   2804: 'Spare_Fault_2804', class No Acknowledgement, trigger "DB302_HMI_Faults_Carrier43_Faults_3" bit 3
   2805: 'Spare_Fault_2805', class No Acknowledgement, trigger "DB302_HMI_Faults_Carrier43_Faults_3" bit 4
   2806: 'Spare_Fault_2806', class No Acknowledgement, trigger "DB302_HMI_Faults_Carrier43_Faults_3" bit 5
   2807: 'Spare_Fault_2807', class No Acknowledgement, trigger "DB302_HMI_Faults_Carrier43_Faults_3" bit 6
   2808: 'Spare_Fault_2808', class No Acknowledgement, trigger "DB302_HMI_Faults_Carrier43_Faults_3" bit 7
   2809: 'Spare_Fault_2809', class No Acknowledgement, trigger "DB302_HMI_Faults_Carrier43_Faults_3" bit 8
   2810: 'Spare_Fault_2810', class No Acknowledgement, trigger "DB302_HMI_Faults_Carrier43_Faults_3" bit 9
   2811: 'Spare_Fault_2811', class No Acknowledgement, trigger "DB302_HMI_Faults_Carrier43_Faults_3" bit 10
   2812: 'Spare_Fault_2812', class No Acknowledgement, trigger "DB302_HMI_Faults_Carrier43_Faults_3" bit 11
   2813: 'Spare_Fault_2813', class No Acknowledgement, trigger "DB302_HMI_Faults_Carrier43_Faults_3" bit 12
   2814: 'Spare_Fault_2814', class No Acknowledgement, trigger "DB302_HMI_Faults_Carrier43_Faults_3" bit 13
   2815: 'Spare_Fault_2815', class No Acknowledgement, trigger "DB302_HMI_Faults_Carrier43_Faults_3" bit 14
   2816: 'Spare_Fault_2816', class No Acknowledgement, trigger "DB302_HMI_Faults_Carrier43_Faults_3" bit 15
   2817: 'Carrier 44 Disconnect Open Power Fault DI11.0', class No Acknowledgement, trigger "DB302_HMI_Faults_Carrier44_Faults_0" bit 0
   2818: 'Carrier 44 Drive Profinet Comm Fault', class No Acknowledgement, trigger "DB302_HMI_Faults_Carrier44_Faults_0" bit 1
   2819: 'Carrier 44 Production Stop Not Reset', class No Acknowledgement, trigger "DB302_HMI_Faults_Carrier44_Faults_0" bit 2
   2820: 'Carrier 44 CB02122 Tripped', class No Acknowledgement, trigger "DB302_HMI_Faults_Carrier44_Faults_0" bit 3
   2821: 'Carrier 44 CB02123 Tripped', class No Acknowledgement, trigger "DB302_HMI_Faults_Carrier44_Faults_0" bit 4
   2822: 'Carrier 44 AUX1 CB Tripped', class No Acknowledgement, trigger "DB302_HMI_Faults_Carrier44_Faults_0" bit 5
   2823: 'Carrier 44 AUX2 CB Tripped', class No Acknowledgement, trigger "DB302_HMI_Faults_Carrier44_Faults_0" bit 6
   2824: 'Carrier 44 PLC Not Communicating', class No Acknowledgement, trigger "DB302_HMI_Faults_Carrier44_Faults_0" bit 7
   2825: 'Carrier 44 Safe Input Card Fault', class No Acknowledgement, trigger "DB302_HMI_Faults_Carrier44_Faults_0" bit 8
   2826: 'Carrier 44 Safe Output Card Fault', class No Acknowledgement, trigger "DB302_HMI_Faults_Carrier44_Faults_0" bit 9
   2827: 'Carrier 44 Standard Input Card Fault', class No Acknowledgement, trigger "DB302_HMI_Faults_Carrier44_Faults_0" bit 10
   2828: 'Carrier 44 Standard Output Card Fault', class No Acknowledgement, trigger "DB302_HMI_Faults_Carrier44_Faults_0" bit 11
   2829: 'Carrier 44 Encoder Position Fault', class No Acknowledgement, trigger "DB302_HMI_Faults_Carrier44_Faults_0" bit 12
   2830: 'Carrier 44 Encoder Internal Error', class No Acknowledgement, trigger "DB302_HMI_Faults_Carrier44_Faults_0" bit 13
   2831: 'Carrier 44 Encoder Comm Fault', class No Acknowledgement, trigger "DB302_HMI_Faults_Carrier44_Faults_0" bit 14
   2832: 'Carrier 44 HMI Comm Fault', class No Acknowledgement, trigger "DB302_HMI_Faults_Carrier44_Faults_0" bit 15
   2833: 'Carrier 44 Crash Detection Fault', class No Acknowledgement, trigger "DB302_HMI_Faults_Carrier44_Faults_1" bit 0
   2834: 'Carrier 44 Carrier Number Invalid', class No Acknowledgement, trigger "DB302_HMI_Faults_Carrier44_Faults_1" bit 1
   2835: 'Carrier 44 Drive: PROFINET configuration error', class No Acknowledgement, trigger "DB302_HMI_Faults_Carrier44_Faults_1" bit 2
   2836: 'Carrier 44 Drive: Error internal communications', class No Acknowledgement, trigger "DB302_HMI_Faults_Carrier44_Faults_1" bit 3
   2837: 'Carrier 44 Drive: Motor overtemperature', class No Acknowledgement, trigger "DB302_HMI_Faults_Carrier44_Faults_1" bit 4
   2838: 'Carrier 44 Drive: Motor overcurrent', class No Acknowledgement, trigger "DB302_HMI_Faults_Carrier44_Faults_1" bit 5
   2839: 'Carrier 44 Drive: Infeed or power unit not ready', class No Acknowledgement, trigger "DB302_HMI_Faults_Carrier44_Faults_1" bit 6
   2840: 'Carrier 44 Drive: Short-circuit/ground fault detected', class No Acknowledgement, trigger "DB302_HMI_Faults_Carrier44_Faults_1" bit 7
   2841: 'Carrier 44 Drive: PROFINET Setpoint timeout', class No Acknowledgement, trigger "DB302_HMI_Faults_Carrier44_Faults_1" bit 8
   2842: 'Carrier 44 Power unit: Overcurrent', class No Acknowledgement, trigger "DB302_HMI_Faults_Carrier44_Faults_1" bit 9
   2843: 'Carrier 44 Power unit: DC link voltage overvoltage', class No Acknowledgement, trigger "DB302_HMI_Faults_Carrier44_Faults_1" bit 10
   2844: 'Carrier 44 Power unit: DC link voltage undervoltage', class No Acknowledgement, trigger "DB302_HMI_Faults_Carrier44_Faults_1" bit 11
   2845: 'Carrier 44 Power unit: Line phase failure in main circuit', class No Acknowledgement, trigger "DB302_HMI_Faults_Carrier44_Faults_1" bit 12
   2846: 'Carrier 44 Power unit: Phase failure motor cable', class No Acknowledgement, trigger "DB302_HMI_Faults_Carrier44_Faults_1" bit 13
   2847: 'Carrier 44 Power unit: Ground fault', class No Acknowledgement, trigger "DB302_HMI_Faults_Carrier44_Faults_1" bit 14
   2848: 'Spare_Fault_2848', class No Acknowledgement, trigger "DB302_HMI_Faults_Carrier44_Faults_1" bit 15
   2849: 'Carrier 44 Motion Off Fault', class No Acknowledgement, trigger "DB302_HMI_Faults_Carrier44_Faults_2" bit 0
   2850: 'Carrier 44 Motion On Fault', class No Acknowledgement, trigger "DB302_HMI_Faults_Carrier44_Faults_2" bit 1
   2851: 'Carrier 44 Spacing Fault', class No Acknowledgement, trigger "DB302_HMI_Faults_Carrier44_Faults_2" bit 2
   2852: 'Carrier 44 Duplicate Carrier Number Fault', class No Acknowledgement, trigger "DB302_HMI_Faults_Carrier44_Faults_2" bit 3
   2853: 'Spare_Fault_2853', class No Acknowledgement, trigger "DB302_HMI_Faults_Carrier44_Faults_2" bit 4
   2854: 'Spare_Fault_2854', class No Acknowledgement, trigger "DB302_HMI_Faults_Carrier44_Faults_2" bit 5
   2855: 'Spare_Fault_2855', class No Acknowledgement, trigger "DB302_HMI_Faults_Carrier44_Faults_2" bit 6
   2856: 'Spare_Fault_2856', class No Acknowledgement, trigger "DB302_HMI_Faults_Carrier44_Faults_2" bit 7
   2857: 'Spare_Fault_2857', class No Acknowledgement, trigger "DB302_HMI_Faults_Carrier44_Faults_2" bit 8
   2858: 'Spare_Fault_2858', class No Acknowledgement, trigger "DB302_HMI_Faults_Carrier44_Faults_2" bit 9
   2859: 'Spare_Fault_2859', class No Acknowledgement, trigger "DB302_HMI_Faults_Carrier44_Faults_2" bit 10
   2860: 'Spare_Fault_2860', class No Acknowledgement, trigger "DB302_HMI_Faults_Carrier44_Faults_2" bit 11
   2861: 'Spare_Fault_2861', class No Acknowledgement, trigger "DB302_HMI_Faults_Carrier44_Faults_2" bit 12
   2862: 'Spare_Fault_2862', class No Acknowledgement, trigger "DB302_HMI_Faults_Carrier44_Faults_2" bit 13
   2863: 'Spare_Fault_2863', class No Acknowledgement, trigger "DB302_HMI_Faults_Carrier44_Faults_2" bit 14
   2864: 'Spare_Fault_2864', class No Acknowledgement, trigger "DB302_HMI_Faults_Carrier44_Faults_2" bit 15
   2865: 'Spare_Fault_2865', class No Acknowledgement, trigger "DB302_HMI_Faults_Carrier44_Faults_3" bit 0
   2866: 'Spare_Fault_2866', class No Acknowledgement, trigger "DB302_HMI_Faults_Carrier44_Faults_3" bit 1
   2867: 'Spare_Fault_2867', class No Acknowledgement, trigger "DB302_HMI_Faults_Carrier44_Faults_3" bit 2
   2868: 'Spare_Fault_2868', class No Acknowledgement, trigger "DB302_HMI_Faults_Carrier44_Faults_3" bit 3
   2869: 'Spare_Fault_2869', class No Acknowledgement, trigger "DB302_HMI_Faults_Carrier44_Faults_3" bit 4
   2870: 'Spare_Fault_2870', class No Acknowledgement, trigger "DB302_HMI_Faults_Carrier44_Faults_3" bit 5
   2871: 'Spare_Fault_2871', class No Acknowledgement, trigger "DB302_HMI_Faults_Carrier44_Faults_3" bit 6
   2872: 'Spare_Fault_2872', class No Acknowledgement, trigger "DB302_HMI_Faults_Carrier44_Faults_3" bit 7
   2873: 'Spare_Fault_2873', class No Acknowledgement, trigger "DB302_HMI_Faults_Carrier44_Faults_3" bit 8
   2874: 'Spare_Fault_2874', class No Acknowledgement, trigger "DB302_HMI_Faults_Carrier44_Faults_3" bit 9
   2875: 'Spare_Fault_2875', class No Acknowledgement, trigger "DB302_HMI_Faults_Carrier44_Faults_3" bit 10
   2876: 'Spare_Fault_2876', class No Acknowledgement, trigger "DB302_HMI_Faults_Carrier44_Faults_3" bit 11
   2877: 'Spare_Fault_2877', class No Acknowledgement, trigger "DB302_HMI_Faults_Carrier44_Faults_3" bit 12
   2878: 'Spare_Fault_2878', class No Acknowledgement, trigger "DB302_HMI_Faults_Carrier44_Faults_3" bit 13
   2879: 'Spare_Fault_2879', class No Acknowledgement, trigger "DB302_HMI_Faults_Carrier44_Faults_3" bit 14
   2880: 'Spare_Fault_2880', class No Acknowledgement, trigger "DB302_HMI_Faults_Carrier44_Faults_3" bit 15
   2881: 'Carrier 45 Disconnect Open Power Fault DI11.0', class No Acknowledgement, trigger "DB302_HMI_Faults_Carrier45_Faults_0" bit 0
   2882: 'Carrier 45 Drive Profinet Comm Fault', class No Acknowledgement, trigger "DB302_HMI_Faults_Carrier45_Faults_0" bit 1
   2883: 'Carrier 45 Production Stop Not Reset', class No Acknowledgement, trigger "DB302_HMI_Faults_Carrier45_Faults_0" bit 2
   2884: 'Carrier 45 CB02122 Tripped', class No Acknowledgement, trigger "DB302_HMI_Faults_Carrier45_Faults_0" bit 3
   2885: 'Carrier 45 CB02123 Tripped', class No Acknowledgement, trigger "DB302_HMI_Faults_Carrier45_Faults_0" bit 4
   2886: 'Carrier 45 AUX1 CB Tripped', class No Acknowledgement, trigger "DB302_HMI_Faults_Carrier45_Faults_0" bit 5
   2887: 'Carrier 45 AUX2 CB Tripped', class No Acknowledgement, trigger "DB302_HMI_Faults_Carrier45_Faults_0" bit 6
   2888: 'Carrier 45 PLC Not Communicating', class No Acknowledgement, trigger "DB302_HMI_Faults_Carrier45_Faults_0" bit 7
   2889: 'Carrier 45 Safe Input Card Fault', class No Acknowledgement, trigger "DB302_HMI_Faults_Carrier45_Faults_0" bit 8
   2890: 'Carrier 45 Safe Output Card Fault', class No Acknowledgement, trigger "DB302_HMI_Faults_Carrier45_Faults_0" bit 9
   2891: 'Carrier 45 Standard Input Card Fault', class No Acknowledgement, trigger "DB302_HMI_Faults_Carrier45_Faults_0" bit 10
   2892: 'Carrier 45 Standard Output Card Fault', class No Acknowledgement, trigger "DB302_HMI_Faults_Carrier45_Faults_0" bit 11
   2893: 'Carrier 45 Encoder Position Fault', class No Acknowledgement, trigger "DB302_HMI_Faults_Carrier45_Faults_0" bit 12
   2894: 'Carrier 45 Encoder Internal Error', class No Acknowledgement, trigger "DB302_HMI_Faults_Carrier45_Faults_0" bit 13
   2895: 'Carrier 45 Encoder Comm Fault', class No Acknowledgement, trigger "DB302_HMI_Faults_Carrier45_Faults_0" bit 14
   2896: 'Carrier 45 HMI Comm Fault', class No Acknowledgement, trigger "DB302_HMI_Faults_Carrier45_Faults_0" bit 15
   2897: 'Carrier 45 Crash Detection Fault', class No Acknowledgement, trigger "DB302_HMI_Faults_Carrier45_Faults_1" bit 0
   2898: 'Carrier 45 Carrier Number Invalid', class No Acknowledgement, trigger "DB302_HMI_Faults_Carrier45_Faults_1" bit 1
   2899: 'Carrier 45 Drive: PROFINET configuration error', class No Acknowledgement, trigger "DB302_HMI_Faults_Carrier45_Faults_1" bit 2
   2900: 'Carrier 45 Drive: Error internal communications', class No Acknowledgement, trigger "DB302_HMI_Faults_Carrier45_Faults_1" bit 3
   2901: 'Carrier 45 Drive: Motor overtemperature', class No Acknowledgement, trigger "DB302_HMI_Faults_Carrier45_Faults_1" bit 4
   2902: 'Carrier 45 Drive: Motor overcurrent', class No Acknowledgement, trigger "DB302_HMI_Faults_Carrier45_Faults_1" bit 5
   2903: 'Carrier 45 Drive: Infeed or power unit not ready', class No Acknowledgement, trigger "DB302_HMI_Faults_Carrier45_Faults_1" bit 6
   2904: 'Carrier 45 Drive: Short-circuit/ground fault detected', class No Acknowledgement, trigger "DB302_HMI_Faults_Carrier45_Faults_1" bit 7
   2905: 'Carrier 45 Drive: PROFINET Setpoint timeout', class No Acknowledgement, trigger "DB302_HMI_Faults_Carrier45_Faults_1" bit 8
   2906: 'Carrier 45 Power unit: Overcurrent', class No Acknowledgement, trigger "DB302_HMI_Faults_Carrier45_Faults_1" bit 9
   2907: 'Carrier 45 Power unit: DC link voltage overvoltage', class No Acknowledgement, trigger "DB302_HMI_Faults_Carrier45_Faults_1" bit 10
   2908: 'Carrier 45 Power unit: DC link voltage undervoltage', class No Acknowledgement, trigger "DB302_HMI_Faults_Carrier45_Faults_1" bit 11
   2909: 'Carrier 45 Power unit: Line phase failure in main circuit', class No Acknowledgement, trigger "DB302_HMI_Faults_Carrier45_Faults_1" bit 12
   2910: 'Carrier 45 Power unit: Phase failure motor cable', class No Acknowledgement, trigger "DB302_HMI_Faults_Carrier45_Faults_1" bit 13
   2911: 'Carrier 45 Power unit: Ground fault', class No Acknowledgement, trigger "DB302_HMI_Faults_Carrier45_Faults_1" bit 14
   2912: 'Spare_Fault_2912', class No Acknowledgement, trigger "DB302_HMI_Faults_Carrier45_Faults_1" bit 15
   2913: 'Carrier 45 Motion Off Fault', class No Acknowledgement, trigger "DB302_HMI_Faults_Carrier45_Faults_2" bit 0
   2914: 'Carrier 45 Motion On Fault', class No Acknowledgement, trigger "DB302_HMI_Faults_Carrier45_Faults_2" bit 1
   2915: 'Carrier 45 Spacing Fault', class No Acknowledgement, trigger "DB302_HMI_Faults_Carrier45_Faults_2" bit 2
   2916: 'Carrier 45 Duplicate Carrier Number Fault', class No Acknowledgement, trigger "DB302_HMI_Faults_Carrier45_Faults_2" bit 3
   2917: 'Spare_Fault_2917', class No Acknowledgement, trigger "DB302_HMI_Faults_Carrier45_Faults_2" bit 4
   2918: 'Spare_Fault_2918', class No Acknowledgement, trigger "DB302_HMI_Faults_Carrier45_Faults_2" bit 5
   2919: 'Spare_Fault_2919', class No Acknowledgement, trigger "DB302_HMI_Faults_Carrier45_Faults_2" bit 6
   2920: 'Spare_Fault_2920', class No Acknowledgement, trigger "DB302_HMI_Faults_Carrier45_Faults_2" bit 7
   2921: 'Spare_Fault_2921', class No Acknowledgement, trigger "DB302_HMI_Faults_Carrier45_Faults_2" bit 8
   2922: 'Spare_Fault_2922', class No Acknowledgement, trigger "DB302_HMI_Faults_Carrier45_Faults_2" bit 9
   2923: 'Spare_Fault_2923', class No Acknowledgement, trigger "DB302_HMI_Faults_Carrier45_Faults_2" bit 10
   2924: 'Spare_Fault_2924', class No Acknowledgement, trigger "DB302_HMI_Faults_Carrier45_Faults_2" bit 11
   2925: 'Spare_Fault_2925', class No Acknowledgement, trigger "DB302_HMI_Faults_Carrier45_Faults_2" bit 12
   2926: 'Spare_Fault_2926', class No Acknowledgement, trigger "DB302_HMI_Faults_Carrier45_Faults_2" bit 13
   2927: 'Spare_Fault_2927', class No Acknowledgement, trigger "DB302_HMI_Faults_Carrier45_Faults_2" bit 14
   2928: 'Spare_Fault_2928', class No Acknowledgement, trigger "DB302_HMI_Faults_Carrier45_Faults_2" bit 15
   2929: 'Spare_Fault_2929', class No Acknowledgement, trigger "DB302_HMI_Faults_Carrier45_Faults_3" bit 0
   2930: 'Spare_Fault_2930', class No Acknowledgement, trigger "DB302_HMI_Faults_Carrier45_Faults_3" bit 1
   2931: 'Spare_Fault_2931', class No Acknowledgement, trigger "DB302_HMI_Faults_Carrier45_Faults_3" bit 2
   2932: 'Spare_Fault_2932', class No Acknowledgement, trigger "DB302_HMI_Faults_Carrier45_Faults_3" bit 3
   2933: 'Spare_Fault_2933', class No Acknowledgement, trigger "DB302_HMI_Faults_Carrier45_Faults_3" bit 4
   2934: 'Spare_Fault_2934', class No Acknowledgement, trigger "DB302_HMI_Faults_Carrier45_Faults_3" bit 5
   2935: 'Spare_Fault_2935', class No Acknowledgement, trigger "DB302_HMI_Faults_Carrier45_Faults_3" bit 6
   2936: 'Spare_Fault_2936', class No Acknowledgement, trigger "DB302_HMI_Faults_Carrier45_Faults_3" bit 7
   2937: 'Spare_Fault_2937', class No Acknowledgement, trigger "DB302_HMI_Faults_Carrier45_Faults_3" bit 8
   2938: 'Spare_Fault_2938', class No Acknowledgement, trigger "DB302_HMI_Faults_Carrier45_Faults_3" bit 9
   2939: 'Spare_Fault_2939', class No Acknowledgement, trigger "DB302_HMI_Faults_Carrier45_Faults_3" bit 10
   2940: 'Spare_Fault_2940', class No Acknowledgement, trigger "DB302_HMI_Faults_Carrier45_Faults_3" bit 11
   2941: 'Spare_Fault_2941', class No Acknowledgement, trigger "DB302_HMI_Faults_Carrier45_Faults_3" bit 12
   2942: 'Spare_Fault_2942', class No Acknowledgement, trigger "DB302_HMI_Faults_Carrier45_Faults_3" bit 13
   2943: 'Spare_Fault_2943', class No Acknowledgement, trigger "DB302_HMI_Faults_Carrier45_Faults_3" bit 14
   2944: 'Spare_Fault_2944', class No Acknowledgement, trigger "DB302_HMI_Faults_Carrier45_Faults_3" bit 15
   2945: 'Carrier 46 Disconnect Open Power Fault DI11.0', class No Acknowledgement, trigger "DB302_HMI_Faults_Carrier46_Faults_0" bit 0
   2946: 'Carrier 46 Drive Profinet Comm Fault', class No Acknowledgement, trigger "DB302_HMI_Faults_Carrier46_Faults_0" bit 1
   2947: 'Carrier 46 Production Stop Not Reset', class No Acknowledgement, trigger "DB302_HMI_Faults_Carrier46_Faults_0" bit 2
   2948: 'Carrier 46 CB02122 Tripped', class No Acknowledgement, trigger "DB302_HMI_Faults_Carrier46_Faults_0" bit 3
   2949: 'Carrier 46 CB02123 Tripped', class No Acknowledgement, trigger "DB302_HMI_Faults_Carrier46_Faults_0" bit 4
   2950: 'Carrier 46 AUX1 CB Tripped', class No Acknowledgement, trigger "DB302_HMI_Faults_Carrier46_Faults_0" bit 5
   2951: 'Carrier 46 AUX2 CB Tripped', class No Acknowledgement, trigger "DB302_HMI_Faults_Carrier46_Faults_0" bit 6
   2952: 'Carrier 46 PLC Not Communicating', class No Acknowledgement, trigger "DB302_HMI_Faults_Carrier46_Faults_0" bit 7
   2953: 'Carrier 46 Safe Input Card Fault', class No Acknowledgement, trigger "DB302_HMI_Faults_Carrier46_Faults_0" bit 8
   2954: 'Carrier 46 Safe Output Card Fault', class No Acknowledgement, trigger "DB302_HMI_Faults_Carrier46_Faults_0" bit 9
   2955: 'Carrier 46 Standard Input Card Fault', class No Acknowledgement, trigger "DB302_HMI_Faults_Carrier46_Faults_0" bit 10
   2956: 'Carrier 46 Standard Output Card Fault', class No Acknowledgement, trigger "DB302_HMI_Faults_Carrier46_Faults_0" bit 11
   2957: 'Carrier 46 Encoder Position Fault', class No Acknowledgement, trigger "DB302_HMI_Faults_Carrier46_Faults_0" bit 12
   2958: 'Carrier 46 Encoder Internal Error', class No Acknowledgement, trigger "DB302_HMI_Faults_Carrier46_Faults_0" bit 13
   2959: 'Carrier 46 Encoder Comm Fault', class No Acknowledgement, trigger "DB302_HMI_Faults_Carrier46_Faults_0" bit 14
   2960: 'Carrier 46 HMI Comm Fault', class No Acknowledgement, trigger "DB302_HMI_Faults_Carrier46_Faults_0" bit 15
   2961: 'Carrier 46 Crash Detection Fault', class No Acknowledgement, trigger "DB302_HMI_Faults_Carrier46_Faults_1" bit 0
   2962: 'Carrier 46 Carrier Number Invalid', class No Acknowledgement, trigger "DB302_HMI_Faults_Carrier46_Faults_1" bit 1
   2963: 'Carrier 46 Drive: PROFINET configuration error', class No Acknowledgement, trigger "DB302_HMI_Faults_Carrier46_Faults_1" bit 2
   2964: 'Carrier 46 Drive: Error internal communications', class No Acknowledgement, trigger "DB302_HMI_Faults_Carrier46_Faults_1" bit 3
   2965: 'Carrier 46 Drive: Motor overtemperature', class No Acknowledgement, trigger "DB302_HMI_Faults_Carrier46_Faults_1" bit 4
   2966: 'Carrier 46 Drive: Motor overcurrent', class No Acknowledgement, trigger "DB302_HMI_Faults_Carrier46_Faults_1" bit 5
   2967: 'Carrier 46 Drive: Infeed or power unit not ready', class No Acknowledgement, trigger "DB302_HMI_Faults_Carrier46_Faults_1" bit 6
   2968: 'Carrier 46 Drive: Short-circuit/ground fault detected', class No Acknowledgement, trigger "DB302_HMI_Faults_Carrier46_Faults_1" bit 7
   2969: 'Carrier 46 Drive: PROFINET Setpoint timeout', class No Acknowledgement, trigger "DB302_HMI_Faults_Carrier46_Faults_1" bit 8
   2970: 'Carrier 46 Power unit: Overcurrent', class No Acknowledgement, trigger "DB302_HMI_Faults_Carrier46_Faults_1" bit 9
   2971: 'Carrier 46 Power unit: DC link voltage overvoltage', class No Acknowledgement, trigger "DB302_HMI_Faults_Carrier46_Faults_1" bit 10
   2972: 'Carrier 46 Power unit: DC link voltage undervoltage', class No Acknowledgement, trigger "DB302_HMI_Faults_Carrier46_Faults_1" bit 11
   2973: 'Carrier 46 Power unit: Line phase failure in main circuit', class No Acknowledgement, trigger "DB302_HMI_Faults_Carrier46_Faults_1" bit 12
   2974: 'Carrier 46 Power unit: Phase failure motor cable', class No Acknowledgement, trigger "DB302_HMI_Faults_Carrier46_Faults_1" bit 13
   2975: 'Carrier 46 Power unit: Ground fault', class No Acknowledgement, trigger "DB302_HMI_Faults_Carrier46_Faults_1" bit 14
   2976: 'Spare_Fault_2976', class No Acknowledgement, trigger "DB302_HMI_Faults_Carrier46_Faults_1" bit 15
   2977: 'Carrier 46 Motion Off Fault', class No Acknowledgement, trigger "DB302_HMI_Faults_Carrier46_Faults_2" bit 0
   2978: 'Carrier 46 Motion On Fault', class No Acknowledgement, trigger "DB302_HMI_Faults_Carrier46_Faults_2" bit 1
   2979: 'Carrier 46 Spacing Fault', class No Acknowledgement, trigger "DB302_HMI_Faults_Carrier46_Faults_2" bit 2
   2980: 'Carrier 46 Duplicate Carrier Number Fault', class No Acknowledgement, trigger "DB302_HMI_Faults_Carrier46_Faults_2" bit 3
   2981: 'Spare_Fault_2981', class No Acknowledgement, trigger "DB302_HMI_Faults_Carrier46_Faults_2" bit 4
   2982: 'Spare_Fault_2982', class No Acknowledgement, trigger "DB302_HMI_Faults_Carrier46_Faults_2" bit 5
   2983: 'Spare_Fault_2983', class No Acknowledgement, trigger "DB302_HMI_Faults_Carrier46_Faults_2" bit 6
   2984: 'Spare_Fault_2984', class No Acknowledgement, trigger "DB302_HMI_Faults_Carrier46_Faults_2" bit 7
   2985: 'Spare_Fault_2985', class No Acknowledgement, trigger "DB302_HMI_Faults_Carrier46_Faults_2" bit 8
   2986: 'Spare_Fault_2986', class No Acknowledgement, trigger "DB302_HMI_Faults_Carrier46_Faults_2" bit 9
   2987: 'Spare_Fault_2987', class No Acknowledgement, trigger "DB302_HMI_Faults_Carrier46_Faults_2" bit 10
   2988: 'Spare_Fault_2988', class No Acknowledgement, trigger "DB302_HMI_Faults_Carrier46_Faults_2" bit 11
   2989: 'Spare_Fault_2989', class No Acknowledgement, trigger "DB302_HMI_Faults_Carrier46_Faults_2" bit 12
   2990: 'Spare_Fault_2990', class No Acknowledgement, trigger "DB302_HMI_Faults_Carrier46_Faults_2" bit 13
   2991: 'Spare_Fault_2991', class No Acknowledgement, trigger "DB302_HMI_Faults_Carrier46_Faults_2" bit 14
   2992: 'Spare_Fault_2992', class No Acknowledgement, trigger "DB302_HMI_Faults_Carrier46_Faults_2" bit 15
   2993: 'Spare_Fault_2993', class No Acknowledgement, trigger "DB302_HMI_Faults_Carrier46_Faults_3" bit 0
   2994: 'Spare_Fault_2994', class No Acknowledgement, trigger "DB302_HMI_Faults_Carrier46_Faults_3" bit 1
   2995: 'Spare_Fault_2995', class No Acknowledgement, trigger "DB302_HMI_Faults_Carrier46_Faults_3" bit 2
   2996: 'Spare_Fault_2996', class No Acknowledgement, trigger "DB302_HMI_Faults_Carrier46_Faults_3" bit 3
   2997: 'Spare_Fault_2997', class No Acknowledgement, trigger "DB302_HMI_Faults_Carrier46_Faults_3" bit 4
   2998: 'Spare_Fault_2998', class No Acknowledgement, trigger "DB302_HMI_Faults_Carrier46_Faults_3" bit 5
   2999: 'Spare_Fault_2999', class No Acknowledgement, trigger "DB302_HMI_Faults_Carrier46_Faults_3" bit 6
   3000: 'Spare_Fault_3000', class No Acknowledgement, trigger "DB302_HMI_Faults_Carrier46_Faults_3" bit 7
   3001: 'Spare_Fault_3001', class No Acknowledgement, trigger "DB302_HMI_Faults_Carrier46_Faults_3" bit 8
   3002: 'Spare_Fault_3002', class No Acknowledgement, trigger "DB302_HMI_Faults_Carrier46_Faults_3" bit 9
   3003: 'Spare_Fault_3003', class No Acknowledgement, trigger "DB302_HMI_Faults_Carrier46_Faults_3" bit 10
   3004: 'Spare_Fault_3004', class No Acknowledgement, trigger "DB302_HMI_Faults_Carrier46_Faults_3" bit 11
   3005: 'Spare_Fault_3005', class No Acknowledgement, trigger "DB302_HMI_Faults_Carrier46_Faults_3" bit 12
   3006: 'Spare_Fault_3006', class No Acknowledgement, trigger "DB302_HMI_Faults_Carrier46_Faults_3" bit 13
   3007: 'Spare_Fault_3007', class No Acknowledgement, trigger "DB302_HMI_Faults_Carrier46_Faults_3" bit 14
   3008: 'Spare_Fault_3008', class No Acknowledgement, trigger "DB302_HMI_Faults_Carrier46_Faults_3" bit 15
   3009: 'Carrier 47 Disconnect Open Power Fault DI11.0', class No Acknowledgement, trigger "DB302_HMI_Faults_Carrier47_Faults_0" bit 0
   3010: 'Carrier 47 Drive Profinet Comm Fault', class No Acknowledgement, trigger "DB302_HMI_Faults_Carrier47_Faults_0" bit 1
   3011: 'Carrier 47 Production Stop Not Reset', class No Acknowledgement, trigger "DB302_HMI_Faults_Carrier47_Faults_0" bit 2
   3012: 'Carrier 47 CB02122 Tripped', class No Acknowledgement, trigger "DB302_HMI_Faults_Carrier47_Faults_0" bit 3
   3013: 'Carrier 47 CB02123 Tripped', class No Acknowledgement, trigger "DB302_HMI_Faults_Carrier47_Faults_0" bit 4
   3014: 'Carrier 47 AUX1 CB Tripped', class No Acknowledgement, trigger "DB302_HMI_Faults_Carrier47_Faults_0" bit 5
   3015: 'Carrier 47 AUX2 CB Tripped', class No Acknowledgement, trigger "DB302_HMI_Faults_Carrier47_Faults_0" bit 6
   3016: 'Carrier 47 PLC Not Communicating', class No Acknowledgement, trigger "DB302_HMI_Faults_Carrier47_Faults_0" bit 7
   3017: 'Carrier 47 Safe Input Card Fault', class No Acknowledgement, trigger "DB302_HMI_Faults_Carrier47_Faults_0" bit 8
   3018: 'Carrier 47 Safe Output Card Fault', class No Acknowledgement, trigger "DB302_HMI_Faults_Carrier47_Faults_0" bit 9
   3019: 'Carrier 47 Standard Input Card Fault', class No Acknowledgement, trigger "DB302_HMI_Faults_Carrier47_Faults_0" bit 10
   3020: 'Carrier 47 Standard Output Card Fault', class No Acknowledgement, trigger "DB302_HMI_Faults_Carrier47_Faults_0" bit 11
   3021: 'Carrier 47 Encoder Position Fault', class No Acknowledgement, trigger "DB302_HMI_Faults_Carrier47_Faults_0" bit 12
   3022: 'Carrier 47 Encoder Internal Error', class No Acknowledgement, trigger "DB302_HMI_Faults_Carrier47_Faults_0" bit 13
   3023: 'Carrier 47 Encoder Comm Fault', class No Acknowledgement, trigger "DB302_HMI_Faults_Carrier47_Faults_0" bit 14
   3024: 'Carrier 47 HMI Comm Fault', class No Acknowledgement, trigger "DB302_HMI_Faults_Carrier47_Faults_0" bit 15
   3025: 'Carrier 47 Crash Detection Fault', class No Acknowledgement, trigger "DB302_HMI_Faults_Carrier47_Faults_1" bit 0
   3026: 'Carrier 47 Carrier Number Invalid', class No Acknowledgement, trigger "DB302_HMI_Faults_Carrier47_Faults_1" bit 1
   3027: 'Carrier 47 Drive: PROFINET configuration error', class No Acknowledgement, trigger "DB302_HMI_Faults_Carrier47_Faults_1" bit 2
   3028: 'Carrier 47 Drive: Error internal communications', class No Acknowledgement, trigger "DB302_HMI_Faults_Carrier47_Faults_1" bit 3
   3029: 'Carrier 47 Drive: Motor overtemperature', class No Acknowledgement, trigger "DB302_HMI_Faults_Carrier47_Faults_1" bit 4
   3030: 'Carrier 47 Drive: Motor overcurrent', class No Acknowledgement, trigger "DB302_HMI_Faults_Carrier47_Faults_1" bit 5
   3031: 'Carrier 47 Drive: Infeed or power unit not ready', class No Acknowledgement, trigger "DB302_HMI_Faults_Carrier47_Faults_1" bit 6
   3032: 'Carrier 47 Drive: Short-circuit/ground fault detected', class No Acknowledgement, trigger "DB302_HMI_Faults_Carrier47_Faults_1" bit 7
   3033: 'Carrier 47 Drive: PROFINET Setpoint timeout', class No Acknowledgement, trigger "DB302_HMI_Faults_Carrier47_Faults_1" bit 8
   3034: 'Carrier 47 Power unit: Overcurrent', class No Acknowledgement, trigger "DB302_HMI_Faults_Carrier47_Faults_1" bit 9
   3035: 'Carrier 47 Power unit: DC link voltage overvoltage', class No Acknowledgement, trigger "DB302_HMI_Faults_Carrier47_Faults_1" bit 10
   3036: 'Carrier 47 Power unit: DC link voltage undervoltage', class No Acknowledgement, trigger "DB302_HMI_Faults_Carrier47_Faults_1" bit 11
   3037: 'Carrier 47 Power unit: Line phase failure in main circuit', class No Acknowledgement, trigger "DB302_HMI_Faults_Carrier47_Faults_1" bit 12
   3038: 'Carrier 47 Power unit: Phase failure motor cable', class No Acknowledgement, trigger "DB302_HMI_Faults_Carrier47_Faults_1" bit 13
   3039: 'Carrier 47 Power unit: Ground fault', class No Acknowledgement, trigger "DB302_HMI_Faults_Carrier47_Faults_1" bit 14
   3040: 'Spare_Fault_3040', class No Acknowledgement, trigger "DB302_HMI_Faults_Carrier47_Faults_1" bit 15
   3041: 'Carrier 47 Motion Off Fault', class No Acknowledgement, trigger "DB302_HMI_Faults_Carrier47_Faults_2" bit 0
   3042: 'Carrier 47 Motion On Fault', class No Acknowledgement, trigger "DB302_HMI_Faults_Carrier47_Faults_2" bit 1
   3043: 'Carrier 47 Spacing Fault', class No Acknowledgement, trigger "DB302_HMI_Faults_Carrier47_Faults_2" bit 2
   3044: 'Carrier 47 Duplicate Carrier Number Fault', class No Acknowledgement, trigger "DB302_HMI_Faults_Carrier47_Faults_2" bit 3
   3045: 'Spare_Fault_3045', class No Acknowledgement, trigger "DB302_HMI_Faults_Carrier47_Faults_2" bit 4
   3046: 'Spare_Fault_3046', class No Acknowledgement, trigger "DB302_HMI_Faults_Carrier47_Faults_2" bit 5
   3047: 'Spare_Fault_3047', class No Acknowledgement, trigger "DB302_HMI_Faults_Carrier47_Faults_2" bit 6
   3048: 'Spare_Fault_3048', class No Acknowledgement, trigger "DB302_HMI_Faults_Carrier47_Faults_2" bit 7
   3049: 'Spare_Fault_3049', class No Acknowledgement, trigger "DB302_HMI_Faults_Carrier47_Faults_2" bit 8
   3050: 'Spare_Fault_3050', class No Acknowledgement, trigger "DB302_HMI_Faults_Carrier47_Faults_2" bit 9
   3051: 'Spare_Fault_3051', class No Acknowledgement, trigger "DB302_HMI_Faults_Carrier47_Faults_2" bit 10
   3052: 'Spare_Fault_3052', class No Acknowledgement, trigger "DB302_HMI_Faults_Carrier47_Faults_2" bit 11
   3053: 'Spare_Fault_3053', class No Acknowledgement, trigger "DB302_HMI_Faults_Carrier47_Faults_2" bit 12
   3054: 'Spare_Fault_3054', class No Acknowledgement, trigger "DB302_HMI_Faults_Carrier47_Faults_2" bit 13
   3055: 'Spare_Fault_3055', class No Acknowledgement, trigger "DB302_HMI_Faults_Carrier47_Faults_2" bit 14
   3056: 'Spare_Fault_3056', class No Acknowledgement, trigger "DB302_HMI_Faults_Carrier47_Faults_2" bit 15
   3057: 'Spare_Fault_3057', class No Acknowledgement, trigger "DB302_HMI_Faults_Carrier47_Faults_3" bit 0
   3058: 'Spare_Fault_3058', class No Acknowledgement, trigger "DB302_HMI_Faults_Carrier47_Faults_3" bit 1
   3059: 'Spare_Fault_3059', class No Acknowledgement, trigger "DB302_HMI_Faults_Carrier47_Faults_3" bit 2
   3060: 'Spare_Fault_3060', class No Acknowledgement, trigger "DB302_HMI_Faults_Carrier47_Faults_3" bit 3
   3061: 'Spare_Fault_3061', class No Acknowledgement, trigger "DB302_HMI_Faults_Carrier47_Faults_3" bit 4
   3062: 'Spare_Fault_3062', class No Acknowledgement, trigger "DB302_HMI_Faults_Carrier47_Faults_3" bit 5
   3063: 'Spare_Fault_3063', class No Acknowledgement, trigger "DB302_HMI_Faults_Carrier47_Faults_3" bit 6
   3064: 'Spare_Fault_3064', class No Acknowledgement, trigger "DB302_HMI_Faults_Carrier47_Faults_3" bit 7
   3065: 'Spare_Fault_3065', class No Acknowledgement, trigger "DB302_HMI_Faults_Carrier47_Faults_3" bit 8
   3066: 'Spare_Fault_3066', class No Acknowledgement, trigger "DB302_HMI_Faults_Carrier47_Faults_3" bit 9
   3067: 'Spare_Fault_3067', class No Acknowledgement, trigger "DB302_HMI_Faults_Carrier47_Faults_3" bit 10
   3068: 'Spare_Fault_3068', class No Acknowledgement, trigger "DB302_HMI_Faults_Carrier47_Faults_3" bit 11
   3069: 'Spare_Fault_3069', class No Acknowledgement, trigger "DB302_HMI_Faults_Carrier47_Faults_3" bit 12
   3070: 'Spare_Fault_3070', class No Acknowledgement, trigger "DB302_HMI_Faults_Carrier47_Faults_3" bit 13
   3071: 'Spare_Fault_3071', class No Acknowledgement, trigger "DB302_HMI_Faults_Carrier47_Faults_3" bit 14
   3072: 'Spare_Fault_3072', class No Acknowledgement, trigger "DB302_HMI_Faults_Carrier47_Faults_3" bit 15
   3073: 'Carrier 48 Disconnect Open Power Fault DI11.0', class No Acknowledgement, trigger "DB302_HMI_Faults_Carrier48_Faults_0" bit 0
   3074: 'Carrier 48 Drive Profinet Comm Fault', class No Acknowledgement, trigger "DB302_HMI_Faults_Carrier48_Faults_0" bit 1
   3075: 'Carrier 48 Production Stop Not Reset', class No Acknowledgement, trigger "DB302_HMI_Faults_Carrier48_Faults_0" bit 2
   3076: 'Carrier 48 CB02122 Tripped', class No Acknowledgement, trigger "DB302_HMI_Faults_Carrier48_Faults_0" bit 3
   3077: 'Carrier 48 CB02123 Tripped', class No Acknowledgement, trigger "DB302_HMI_Faults_Carrier48_Faults_0" bit 4
   3078: 'Carrier 48 AUX1 CB Tripped', class No Acknowledgement, trigger "DB302_HMI_Faults_Carrier48_Faults_0" bit 5
   3079: 'Carrier 48 AUX2 CB Tripped', class No Acknowledgement, trigger "DB302_HMI_Faults_Carrier48_Faults_0" bit 6
   3080: 'Carrier 48 PLC Not Communicating', class No Acknowledgement, trigger "DB302_HMI_Faults_Carrier48_Faults_0" bit 7
   3081: 'Carrier 48 Safe Input Card Fault', class No Acknowledgement, trigger "DB302_HMI_Faults_Carrier48_Faults_0" bit 8
   3082: 'Carrier 48 Safe Output Card Fault', class No Acknowledgement, trigger "DB302_HMI_Faults_Carrier48_Faults_0" bit 9
   3083: 'Carrier 48 Standard Input Card Fault', class No Acknowledgement, trigger "DB302_HMI_Faults_Carrier48_Faults_0" bit 10
   3084: 'Carrier 48 Standard Output Card Fault', class No Acknowledgement, trigger "DB302_HMI_Faults_Carrier48_Faults_0" bit 11
   3085: 'Carrier 48 Encoder Position Fault', class No Acknowledgement, trigger "DB302_HMI_Faults_Carrier48_Faults_0" bit 12
   3086: 'Carrier 48 Encoder Internal Error', class No Acknowledgement, trigger "DB302_HMI_Faults_Carrier48_Faults_0" bit 13
   3087: 'Carrier 48 Encoder Comm Fault', class No Acknowledgement, trigger "DB302_HMI_Faults_Carrier48_Faults_0" bit 14
   3088: 'Carrier 48 HMI Comm Fault', class No Acknowledgement, trigger "DB302_HMI_Faults_Carrier48_Faults_0" bit 15
   3089: 'Carrier 48 Crash Detection Fault', class No Acknowledgement, trigger "DB302_HMI_Faults_Carrier48_Faults_1" bit 0
   3090: 'Carrier 48 Carrier Number Invalid', class No Acknowledgement, trigger "DB302_HMI_Faults_Carrier48_Faults_1" bit 1
   3091: 'Carrier 48 Drive: PROFINET configuration error', class No Acknowledgement, trigger "DB302_HMI_Faults_Carrier48_Faults_1" bit 2
   3092: 'Carrier 48 Drive: Error internal communications', class No Acknowledgement, trigger "DB302_HMI_Faults_Carrier48_Faults_1" bit 3
   3093: 'Carrier 48 Drive: Motor overtemperature', class No Acknowledgement, trigger "DB302_HMI_Faults_Carrier48_Faults_1" bit 4
   3094: 'Carrier 48 Drive: Motor overcurrent', class No Acknowledgement, trigger "DB302_HMI_Faults_Carrier48_Faults_1" bit 5
   3095: 'Carrier 48 Drive: Infeed or power unit not ready', class No Acknowledgement, trigger "DB302_HMI_Faults_Carrier48_Faults_1" bit 6
   3096: 'Carrier 48 Drive: Short-circuit/ground fault detected', class No Acknowledgement, trigger "DB302_HMI_Faults_Carrier48_Faults_1" bit 7
   3097: 'Carrier 48 Drive: PROFINET Setpoint timeout', class No Acknowledgement, trigger "DB302_HMI_Faults_Carrier48_Faults_1" bit 8
   3098: 'Carrier 48 Power unit: Overcurrent', class No Acknowledgement, trigger "DB302_HMI_Faults_Carrier48_Faults_1" bit 9
   3099: 'Carrier 48 Power unit: DC link voltage overvoltage', class No Acknowledgement, trigger "DB302_HMI_Faults_Carrier48_Faults_1" bit 10
   3100: 'Carrier 48 Power unit: DC link voltage undervoltage', class No Acknowledgement, trigger "DB302_HMI_Faults_Carrier48_Faults_1" bit 11
   3101: 'Carrier 48 Power unit: Line phase failure in main circuit', class No Acknowledgement, trigger "DB302_HMI_Faults_Carrier48_Faults_1" bit 12
   3102: 'Carrier 48 Power unit: Phase failure motor cable', class No Acknowledgement, trigger "DB302_HMI_Faults_Carrier48_Faults_1" bit 13
   3103: 'Carrier 48 Power unit: Ground fault', class No Acknowledgement, trigger "DB302_HMI_Faults_Carrier48_Faults_1" bit 14
   3104: 'Spare_Fault_3104', class No Acknowledgement, trigger "DB302_HMI_Faults_Carrier48_Faults_1" bit 15
   3105: 'Carrier 48 Motion Off Fault', class No Acknowledgement, trigger "DB302_HMI_Faults_Carrier48_Faults_2" bit 0
   3106: 'Carrier 48 Motion On Fault', class No Acknowledgement, trigger "DB302_HMI_Faults_Carrier48_Faults_2" bit 1
   3107: 'Carrier 48 Spacing Fault', class No Acknowledgement, trigger "DB302_HMI_Faults_Carrier48_Faults_2" bit 2
   3108: 'Carrier 48 Duplicate Carrier Number Fault', class No Acknowledgement, trigger "DB302_HMI_Faults_Carrier48_Faults_2" bit 3
   3109: 'Spare_Fault_3109', class No Acknowledgement, trigger "DB302_HMI_Faults_Carrier48_Faults_2" bit 4
   3110: 'Spare_Fault_3110', class No Acknowledgement, trigger "DB302_HMI_Faults_Carrier48_Faults_2" bit 5
   3111: 'Spare_Fault_3111', class No Acknowledgement, trigger "DB302_HMI_Faults_Carrier48_Faults_2" bit 6
   3112: 'Spare_Fault_3112', class No Acknowledgement, trigger "DB302_HMI_Faults_Carrier48_Faults_2" bit 7
   3113: 'Spare_Fault_3113', class No Acknowledgement, trigger "DB302_HMI_Faults_Carrier48_Faults_2" bit 8
   3114: 'Spare_Fault_3114', class No Acknowledgement, trigger "DB302_HMI_Faults_Carrier48_Faults_2" bit 9
   3115: 'Spare_Fault_3115', class No Acknowledgement, trigger "DB302_HMI_Faults_Carrier48_Faults_2" bit 10
   3116: 'Spare_Fault_3116', class No Acknowledgement, trigger "DB302_HMI_Faults_Carrier48_Faults_2" bit 11
   3117: 'Spare_Fault_3117', class No Acknowledgement, trigger "DB302_HMI_Faults_Carrier48_Faults_2" bit 12
   3118: 'Spare_Fault_3118', class No Acknowledgement, trigger "DB302_HMI_Faults_Carrier48_Faults_2" bit 13
   3119: 'Spare_Fault_3119', class No Acknowledgement, trigger "DB302_HMI_Faults_Carrier48_Faults_2" bit 14
   3120: 'Spare_Fault_3120', class No Acknowledgement, trigger "DB302_HMI_Faults_Carrier48_Faults_2" bit 15
   3121: 'Spare_Fault_3121', class No Acknowledgement, trigger "DB302_HMI_Faults_Carrier48_Faults_3" bit 0
   3122: 'Spare_Fault_3122', class No Acknowledgement, trigger "DB302_HMI_Faults_Carrier48_Faults_3" bit 1
   3123: 'Spare_Fault_3123', class No Acknowledgement, trigger "DB302_HMI_Faults_Carrier48_Faults_3" bit 2
   3124: 'Spare_Fault_3124', class No Acknowledgement, trigger "DB302_HMI_Faults_Carrier48_Faults_3" bit 3
   3125: 'Spare_Fault_3125', class No Acknowledgement, trigger "DB302_HMI_Faults_Carrier48_Faults_3" bit 4
   3126: 'Spare_Fault_3126', class No Acknowledgement, trigger "DB302_HMI_Faults_Carrier48_Faults_3" bit 5
   3127: 'Spare_Fault_3127', class No Acknowledgement, trigger "DB302_HMI_Faults_Carrier48_Faults_3" bit 6
   3128: 'Spare_Fault_3128', class No Acknowledgement, trigger "DB302_HMI_Faults_Carrier48_Faults_3" bit 7
   3129: 'Spare_Fault_3129', class No Acknowledgement, trigger "DB302_HMI_Faults_Carrier48_Faults_3" bit 8
   3130: 'Spare_Fault_3130', class No Acknowledgement, trigger "DB302_HMI_Faults_Carrier48_Faults_3" bit 9
   3131: 'Spare_Fault_3131', class No Acknowledgement, trigger "DB302_HMI_Faults_Carrier48_Faults_3" bit 10
   3132: 'Spare_Fault_3132', class No Acknowledgement, trigger "DB302_HMI_Faults_Carrier48_Faults_3" bit 11
   3133: 'Spare_Fault_3133', class No Acknowledgement, trigger "DB302_HMI_Faults_Carrier48_Faults_3" bit 12
   3134: 'Spare_Fault_3134', class No Acknowledgement, trigger "DB302_HMI_Faults_Carrier48_Faults_3" bit 13
   3135: 'Spare_Fault_3135', class No Acknowledgement, trigger "DB302_HMI_Faults_Carrier48_Faults_3" bit 14
   3136: 'Spare_Fault_3136', class No Acknowledgement, trigger "DB302_HMI_Faults_Carrier48_Faults_3" bit 15
   3137: 'Carrier 49 Disconnect Open Power Fault DI11.0', class No Acknowledgement, trigger "DB302_HMI_Faults_Carrier49_Faults_0" bit 0
   3138: 'Carrier 49 Drive Profinet Comm Fault', class No Acknowledgement, trigger "DB302_HMI_Faults_Carrier49_Faults_0" bit 1
   3139: 'Carrier 49 Production Stop Not Reset', class No Acknowledgement, trigger "DB302_HMI_Faults_Carrier49_Faults_0" bit 2
   3140: 'Carrier 49 CB02122 Tripped', class No Acknowledgement, trigger "DB302_HMI_Faults_Carrier49_Faults_0" bit 3
   3141: 'Carrier 49 CB02123 Tripped', class No Acknowledgement, trigger "DB302_HMI_Faults_Carrier49_Faults_0" bit 4
   3142: 'Carrier 49 AUX1 CB Tripped', class No Acknowledgement, trigger "DB302_HMI_Faults_Carrier49_Faults_0" bit 5
   3143: 'Carrier 49 AUX2 CB Tripped', class No Acknowledgement, trigger "DB302_HMI_Faults_Carrier49_Faults_0" bit 6
   3144: 'Carrier 49 PLC Not Communicating', class No Acknowledgement, trigger "DB302_HMI_Faults_Carrier49_Faults_0" bit 7
   3145: 'Carrier 49 Safe Input Card Fault', class No Acknowledgement, trigger "DB302_HMI_Faults_Carrier49_Faults_0" bit 8
   3146: 'Carrier 49 Safe Output Card Fault', class No Acknowledgement, trigger "DB302_HMI_Faults_Carrier49_Faults_0" bit 9
   3147: 'Carrier 49 Standard Input Card Fault', class No Acknowledgement, trigger "DB302_HMI_Faults_Carrier49_Faults_0" bit 10
   3148: 'Carrier 49 Standard Output Card Fault', class No Acknowledgement, trigger "DB302_HMI_Faults_Carrier49_Faults_0" bit 11
   3149: 'Carrier 49 Encoder Position Fault', class No Acknowledgement, trigger "DB302_HMI_Faults_Carrier49_Faults_0" bit 12
   3150: 'Carrier 49 Encoder Internal Error', class No Acknowledgement, trigger "DB302_HMI_Faults_Carrier49_Faults_0" bit 13
   3151: 'Carrier 49 Encoder Comm Fault', class No Acknowledgement, trigger "DB302_HMI_Faults_Carrier49_Faults_0" bit 14
   3152: 'Carrier 49 HMI Comm Fault', class No Acknowledgement, trigger "DB302_HMI_Faults_Carrier49_Faults_0" bit 15
   3153: 'Carrier 49 Crash Detection Fault', class No Acknowledgement, trigger "DB302_HMI_Faults_Carrier49_Faults_1" bit 0
   3154: 'Carrier 49 Carrier Number Invalid', class No Acknowledgement, trigger "DB302_HMI_Faults_Carrier49_Faults_1" bit 1
   3155: 'Carrier 49 Drive: PROFINET configuration error', class No Acknowledgement, trigger "DB302_HMI_Faults_Carrier49_Faults_1" bit 2
   3156: 'Carrier 49 Drive: Error internal communications', class No Acknowledgement, trigger "DB302_HMI_Faults_Carrier49_Faults_1" bit 3
   3157: 'Carrier 49 Drive: Motor overtemperature', class No Acknowledgement, trigger "DB302_HMI_Faults_Carrier49_Faults_1" bit 4
   3158: 'Carrier 49 Drive: Motor overcurrent', class No Acknowledgement, trigger "DB302_HMI_Faults_Carrier49_Faults_1" bit 5
   3159: 'Carrier 49 Drive: Infeed or power unit not ready', class No Acknowledgement, trigger "DB302_HMI_Faults_Carrier49_Faults_1" bit 6
   3160: 'Carrier 49 Drive: Short-circuit/ground fault detected', class No Acknowledgement, trigger "DB302_HMI_Faults_Carrier49_Faults_1" bit 7
   3161: 'Carrier 49 Drive: PROFINET Setpoint timeout', class No Acknowledgement, trigger "DB302_HMI_Faults_Carrier49_Faults_1" bit 8
   3162: 'Carrier 49 Power unit: Overcurrent', class No Acknowledgement, trigger "DB302_HMI_Faults_Carrier49_Faults_1" bit 9
   3163: 'Carrier 49 Power unit: DC link voltage overvoltage', class No Acknowledgement, trigger "DB302_HMI_Faults_Carrier49_Faults_1" bit 10
   3164: 'Carrier 49 Power unit: DC link voltage undervoltage', class No Acknowledgement, trigger "DB302_HMI_Faults_Carrier49_Faults_1" bit 11
   3165: 'Carrier 49 Power unit: Line phase failure in main circuit', class No Acknowledgement, trigger "DB302_HMI_Faults_Carrier49_Faults_1" bit 12
   3166: 'Carrier 49 Power unit: Phase failure motor cable', class No Acknowledgement, trigger "DB302_HMI_Faults_Carrier49_Faults_1" bit 13
   3167: 'Carrier 49 Power unit: Ground fault', class No Acknowledgement, trigger "DB302_HMI_Faults_Carrier49_Faults_1" bit 14
   3168: 'Spare_Fault_3168', class No Acknowledgement, trigger "DB302_HMI_Faults_Carrier49_Faults_1" bit 15
   3169: 'Carrier 49 Motion Off Fault', class No Acknowledgement, trigger "DB302_HMI_Faults_Carrier49_Faults_2" bit 0
   3170: 'Carrier 49 Motion On Fault', class No Acknowledgement, trigger "DB302_HMI_Faults_Carrier49_Faults_2" bit 1
   3171: 'Carrier 49 Spacing Fault', class No Acknowledgement, trigger "DB302_HMI_Faults_Carrier49_Faults_2" bit 2
   3172: 'Carrier 49 Duplicate Carrier Number Fault', class No Acknowledgement, trigger "DB302_HMI_Faults_Carrier49_Faults_2" bit 3
   3173: 'Spare_Fault_3173', class No Acknowledgement, trigger "DB302_HMI_Faults_Carrier49_Faults_2" bit 4
   3174: 'Spare_Fault_3174', class No Acknowledgement, trigger "DB302_HMI_Faults_Carrier49_Faults_2" bit 5
   3175: 'Spare_Fault_3175', class No Acknowledgement, trigger "DB302_HMI_Faults_Carrier49_Faults_2" bit 6
   3176: 'Spare_Fault_3176', class No Acknowledgement, trigger "DB302_HMI_Faults_Carrier49_Faults_2" bit 7
   3177: 'Spare_Fault_3177', class No Acknowledgement, trigger "DB302_HMI_Faults_Carrier49_Faults_2" bit 8
   3178: 'Spare_Fault_3178', class No Acknowledgement, trigger "DB302_HMI_Faults_Carrier49_Faults_2" bit 9
   3179: 'Spare_Fault_3179', class No Acknowledgement, trigger "DB302_HMI_Faults_Carrier49_Faults_2" bit 10
   3180: 'Spare_Fault_3180', class No Acknowledgement, trigger "DB302_HMI_Faults_Carrier49_Faults_2" bit 11
   3181: 'Spare_Fault_3181', class No Acknowledgement, trigger "DB302_HMI_Faults_Carrier49_Faults_2" bit 12
   3182: 'Spare_Fault_3182', class No Acknowledgement, trigger "DB302_HMI_Faults_Carrier49_Faults_2" bit 13
   3183: 'Spare_Fault_3183', class No Acknowledgement, trigger "DB302_HMI_Faults_Carrier49_Faults_2" bit 14
   3184: 'Spare_Fault_3184', class No Acknowledgement, trigger "DB302_HMI_Faults_Carrier49_Faults_2" bit 15
   3185: 'Spare_Fault_3185', class No Acknowledgement, trigger "DB302_HMI_Faults_Carrier49_Faults_3" bit 0
   3186: 'Spare_Fault_3186', class No Acknowledgement, trigger "DB302_HMI_Faults_Carrier49_Faults_3" bit 1
   3187: 'Spare_Fault_3187', class No Acknowledgement, trigger "DB302_HMI_Faults_Carrier49_Faults_3" bit 2
   3188: 'Spare_Fault_3188', class No Acknowledgement, trigger "DB302_HMI_Faults_Carrier49_Faults_3" bit 3
   3189: 'Spare_Fault_3189', class No Acknowledgement, trigger "DB302_HMI_Faults_Carrier49_Faults_3" bit 4
   3190: 'Spare_Fault_3190', class No Acknowledgement, trigger "DB302_HMI_Faults_Carrier49_Faults_3" bit 5
   3191: 'Spare_Fault_3191', class No Acknowledgement, trigger "DB302_HMI_Faults_Carrier49_Faults_3" bit 6
   3192: 'Spare_Fault_3192', class No Acknowledgement, trigger "DB302_HMI_Faults_Carrier49_Faults_3" bit 7
   3193: 'Spare_Fault_3193', class No Acknowledgement, trigger "DB302_HMI_Faults_Carrier49_Faults_3" bit 8
   3194: 'Spare_Fault_3194', class No Acknowledgement, trigger "DB302_HMI_Faults_Carrier49_Faults_3" bit 9
   3195: 'Spare_Fault_3195', class No Acknowledgement, trigger "DB302_HMI_Faults_Carrier49_Faults_3" bit 10
   3196: 'Spare_Fault_3196', class No Acknowledgement, trigger "DB302_HMI_Faults_Carrier49_Faults_3" bit 11
   3197: 'Spare_Fault_3197', class No Acknowledgement, trigger "DB302_HMI_Faults_Carrier49_Faults_3" bit 12
   3198: 'Spare_Fault_3198', class No Acknowledgement, trigger "DB302_HMI_Faults_Carrier49_Faults_3" bit 13
   3199: 'Spare_Fault_3199', class No Acknowledgement, trigger "DB302_HMI_Faults_Carrier49_Faults_3" bit 14
   3200: 'Spare_Fault_3200', class No Acknowledgement, trigger "DB302_HMI_Faults_Carrier49_Faults_3" bit 15
   3201: 'Carrier 50 Disconnect Open Power Fault DI11.0', class No Acknowledgement, trigger "DB302_HMI_Faults_Carrier50_Faults_0" bit 0
   3202: 'Carrier 50 Drive Profinet Comm Fault', class No Acknowledgement, trigger "DB302_HMI_Faults_Carrier50_Faults_0" bit 1
   3203: 'Carrier 50 Production Stop Not Reset', class No Acknowledgement, trigger "DB302_HMI_Faults_Carrier50_Faults_0" bit 2
   3204: 'Carrier 50 CB02122 Tripped', class No Acknowledgement, trigger "DB302_HMI_Faults_Carrier50_Faults_0" bit 3
   3205: 'Carrier 50 CB02123 Tripped', class No Acknowledgement, trigger "DB302_HMI_Faults_Carrier50_Faults_0" bit 4
   3206: 'Carrier 50 AUX1 CB Tripped', class No Acknowledgement, trigger "DB302_HMI_Faults_Carrier50_Faults_0" bit 5
   3207: 'Carrier 50 AUX2 CB Tripped', class No Acknowledgement, trigger "DB302_HMI_Faults_Carrier50_Faults_0" bit 6
   3208: 'Carrier 50 PLC Not Communicating', class No Acknowledgement, trigger "DB302_HMI_Faults_Carrier50_Faults_0" bit 7
   3209: 'Carrier 50 Safe Input Card Fault', class No Acknowledgement, trigger "DB302_HMI_Faults_Carrier50_Faults_0" bit 8
   3210: 'Carrier 50 Safe Output Card Fault', class No Acknowledgement, trigger "DB302_HMI_Faults_Carrier50_Faults_0" bit 9
   3211: 'Carrier 50 Standard Input Card Fault', class No Acknowledgement, trigger "DB302_HMI_Faults_Carrier50_Faults_0" bit 10
   3212: 'Carrier 50 Standard Output Card Fault', class No Acknowledgement, trigger "DB302_HMI_Faults_Carrier50_Faults_0" bit 11
   3213: 'Carrier 50 Encoder Position Fault', class No Acknowledgement, trigger "DB302_HMI_Faults_Carrier50_Faults_0" bit 12
   3214: 'Carrier 50 Encoder Internal Error', class No Acknowledgement, trigger "DB302_HMI_Faults_Carrier50_Faults_0" bit 13
   3215: 'Carrier 50 Encoder Comm Fault', class No Acknowledgement, trigger "DB302_HMI_Faults_Carrier50_Faults_0" bit 14
   3216: 'Carrier 50 HMI Comm Fault', class No Acknowledgement, trigger "DB302_HMI_Faults_Carrier50_Faults_0" bit 15
   3217: 'Carrier 50 Crash Detection Fault', class No Acknowledgement, trigger "DB302_HMI_Faults_Carrier50_Faults_1" bit 0
   3218: 'Carrier 50 Carrier Number Invalid', class No Acknowledgement, trigger "DB302_HMI_Faults_Carrier50_Faults_1" bit 1
   3219: 'Carrier 50 Drive: PROFINET configuration error', class No Acknowledgement, trigger "DB302_HMI_Faults_Carrier50_Faults_1" bit 2
   3220: 'Carrier 50 Drive: Error internal communications', class No Acknowledgement, trigger "DB302_HMI_Faults_Carrier50_Faults_1" bit 3
   3221: 'Carrier 50 Drive: Motor overtemperature', class No Acknowledgement, trigger "DB302_HMI_Faults_Carrier50_Faults_1" bit 4
   3222: 'Carrier 50 Drive: Motor overcurrent', class No Acknowledgement, trigger "DB302_HMI_Faults_Carrier50_Faults_1" bit 5
   3223: 'Carrier 50 Drive: Infeed or power unit not ready', class No Acknowledgement, trigger "DB302_HMI_Faults_Carrier50_Faults_1" bit 6
   3224: 'Carrier 50 Drive: Short-circuit/ground fault detected', class No Acknowledgement, trigger "DB302_HMI_Faults_Carrier50_Faults_1" bit 7
